// TIA Portal project "StepTimeAnalysis" (V16) (continued)
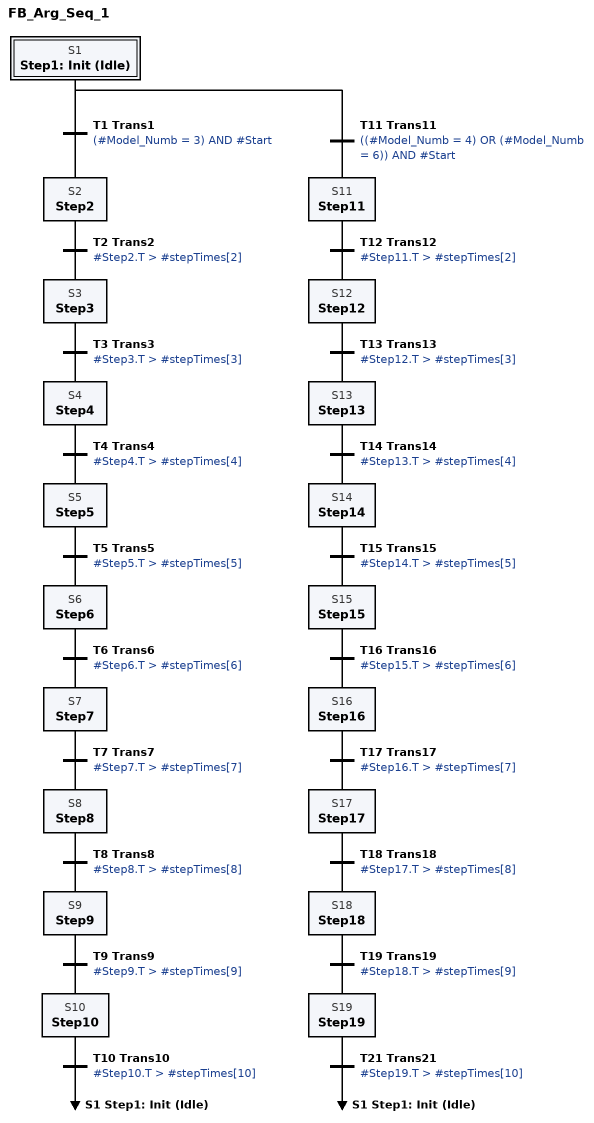
   // sequencer 1
   INITIAL_STEP "Step1: Init (Idle)":   // S1, max time T#10S, warning time T#7S
   END_STEP
   TRANSITION Trans1 FROM "Step1: Init (Idle)" TO Step2   // T1
      := (#Model_Numb = 3) AND #Start;
   END_TRANSITION
   TRANSITION Trans11 FROM "Step1: Init (Idle)" TO Step11   // T11
      := ((#Model_Numb = 4) OR (#Model_Numb = 6)) AND #Start;
   END_TRANSITION
   STEP Step2:   // S2, max time T#10S, warning time T#7S
   END_STEP
   TRANSITION Trans2 FROM Step2 TO Step3   // T2
      := #Step2.T > #stepTimes[2];
   END_TRANSITION
   STEP Step3:   // S3, max time T#10S, warning time T#7S
   END_STEP
   TRANSITION Trans3 FROM Step3 TO Step4   // T3
      := #Step3.T > #stepTimes[3];
   END_TRANSITION
   STEP Step4:   // S4, max time T#10S, warning time T#7S
   END_STEP
   TRANSITION Trans4 FROM Step4 TO Step5   // T4
      := #Step4.T > #stepTimes[4];
   END_TRANSITION
   STEP Step5:   // S5, max time T#10S, warning time T#7S
   END_STEP
   TRANSITION Trans5 FROM Step5 TO Step6   // T5
      := #Step5.T > #stepTimes[5];
   END_TRANSITION
   STEP Step6:   // S6, max time T#10S, warning time T#7S
   END_STEP
   TRANSITION Trans6 FROM Step6 TO Step7   // T6
      := #Step6.T > #stepTimes[6];
   END_TRANSITION
   STEP Step7:   // S7, max time T#10S, warning time T#7S
   END_STEP
   TRANSITION Trans7 FROM Step7 TO Step8   // T7
      := #Step7.T > #stepTimes[7];
   END_TRANSITION
   STEP Step8:   // S8, max time T#10S, warning time T#7S
   END_STEP
   TRANSITION Trans8 FROM Step8 TO Step9   // T8
      := #Step8.T > #stepTimes[8];
   END_TRANSITION
   STEP Step9:   // S9, max time T#10S, warning time T#7S
   END_STEP
   TRANSITION Trans9 FROM Step9 TO Step10   // T9
      := #Step9.T > #stepTimes[9];
   END_TRANSITION
   STEP Step10:   // S10, max time T#10S, warning time T#7S
   END_STEP
   TRANSITION Trans10 FROM Step10 TO "Step1: Init (Idle)"   // T10, jump
      := #Step10.T > #stepTimes[10];
   END_TRANSITION
   STEP Step11:   // S11, max time T#10S, warning time T#7S
   END_STEP
   TRANSITION Trans12 FROM Step11 TO Step12   // T12
      := #Step11.T > #stepTimes[2];
   END_TRANSITION
   STEP Step12:   // S12, max time T#10S, warning time T#7S
   END_STEP
   TRANSITION Trans13 FROM Step12 TO Step13   // T13
      := #Step12.T > #stepTimes[3];
   END_TRANSITION
   STEP Step13:   // S13, max time T#10S, warning time T#7S
   END_STEP
   TRANSITION Trans14 FROM Step13 TO Step14   // T14
      := #Step13.T > #stepTimes[4];
   END_TRANSITION
   STEP Step14:   // S14, max time T#10S, warning time T#7S
   END_STEP
   TRANSITION Trans15 FROM Step14 TO Step15   // T15
      := #Step14.T > #stepTimes[5];
   END_TRANSITION
   STEP Step15:   // S15, max time T#10S, warning time T#7S
   END_STEP
   TRANSITION Trans16 FROM Step15 TO Step16   // T16
      := #Step15.T > #stepTimes[6];
   END_TRANSITION
   STEP Step16:   // S16, max time T#10S, warning time T#7S
   END_STEP
   TRANSITION Trans17 FROM Step16 TO Step17   // T17
      := #Step16.T > #stepTimes[7];
   END_TRANSITION
   STEP Step17:   // S17, max time T#10S, warning time T#7S
   END_STEP
   TRANSITION Trans18 FROM Step17 TO Step18   // T18
      := #Step17.T > #stepTimes[8];
   END_TRANSITION
   STEP Step18:   // S18, max time T#10S, warning time T#7S
   END_STEP
   TRANSITION Trans19 FROM Step18 TO Step19   // T19
      := #Step18.T > #stepTimes[9];
   END_TRANSITION
   STEP Step19:   // S19, max time T#10S, warning time T#7S
   END_STEP
   TRANSITION Trans21 FROM Step19 TO "Step1: Init (Idle)"   // T21, jump
      := #Step19.T > #stepTimes[10];
   END_TRANSITION
END_FUNCTION_BLOCK

FUNCTION "FC_ARG_1" : Void   // FC1, FBD
{ S7_Optimized_Access := 'TRUE' }
VERSION : 0.1
   VAR_OUTPUT
      Ready_new_car : Bool;
   END_VAR
   VAR_TEMP
      stepTimes : Array[2..10] of Time;
      i : Int;
      Random_Time : Time;   // Random Time between 0sec to 10sec
      Start : Bool;
      Stop : Bool;
      status1_RandFunc : Word;
      status2_RandFunc : Word;
      temp : Byte;
      error_RandFunc : Bool;
   END_VAR
   VAR CONSTANT
      sequenceNO : Int := 9;
   END_VAR
BEGIN

REGION Network 1 (SCL): Man Mode Data Handling
   IF "DB_Process_Var".Man_Mode = TRUE THEN
       "DB_Process_Var".Car_Type_Selected := "DB_HMI".dropdown_selection;
   END_IF;
END_REGION

REGION Network 2 (SCL): Auto Mode Data Handling
   IF "DB_Process_Var".Auto_Mode = TRUE THEN
       "DB_HMI".dropdown_selection := 0;
       "DB_Process_Var".Car_Type_Selected := "DB_PLC2_Receiving".ReceivingBoxForward.Type;
   END_IF;
   IF "DB_HMI".ARG1_Seq1_Cmd_Auto OR "DB_HMI".Global_Cmd_Auto THEN
       "DB_HMI".dropdown_selection := 0;
       "DB_Process_Var".Car_Type_Selected := 0;
   END_IF;
END_REGION

REGION Network 3 (SCL): Load Time Date based on Car Type
       CASE "DB_Process_Var".Car_Type_Selected OF
           3:
               "DB_Profile"."time" := "DB_Profile".time_Red;
           4:
               "DB_Profile"."time" := "DB_Profile".time_Green;
           6:
               "DB_Profile"."time" := "DB_Profile".time_Blue;
       END_CASE;
END_REGION

REGION Network 4 (SCL): Switch from selected to inProduction
   IF "IDB_Arg_Seq_1_DB".Trans1.TS = TRUE OR "IDB_Arg_Seq_1_DB".Trans11.TS = TRUE THEN
       IF "DB_Process_Var".Car_Type_Selected = 3 THEN
           "DB_Process_Var".Car_Type_inProduction := 3;
           "DB_Process_Var".Car_Type_inProduction_Text := 'Red';
           "DB_HMI".ARG1_Seq1_inProduction := 3;
       ELSIF "DB_Process_Var".Car_Type_Selected = 4 THEN
           "DB_Process_Var".Car_Type_inProduction := 4;
           "DB_Process_Var".Car_Type_inProduction_Text := 'Green';
           "DB_HMI".ARG1_Seq1_inProduction := 4;
       ELSIF "DB_Process_Var".Car_Type_Selected = 6 THEN
           "DB_Process_Var".Car_Type_inProduction := 6;
           "DB_Process_Var".Car_Type_inProduction_Text := 'Blue';
           "DB_HMI".ARG1_Seq1_inProduction := 6;
       END_IF;
   END_IF;
END_REGION

REGION Network 5 (SCL): Create Random Time Values for the selected Steps
   IF "IDB_Arg_Seq_1_DB".Trans1.TS = TRUE OR "IDB_Arg_Seq_1_DB".Trans11.TS = TRUE THEN
       FOR #i := 2 TO 10 DO
           //Red
           IF "DB_HMI".ARG1_Seq1_DelaySelect_Red[#i] = TRUE THEN;
               "DB_Sim".Delta_T_Red[#i] := "LGF_RandomRange_Dint"(minValue := 0, maxValue := 10000, error => #error_RandFunc, status => #status1_RandFunc, subfunctionStatus => #status2_RandFunc);
           ELSE
               "DB_Sim".Delta_T_Red[#i] := T#0s;
           END_IF;
           //Green
           IF "DB_HMI".ARG1_Seq1_DelaySelect_Green[#i] = TRUE THEN
               "DB_Sim".Delta_T_Green[#i] := "LGF_RandomRange_Dint"(minValue := 0, maxValue := 10000, error => #error_RandFunc, status => #status1_RandFunc, subfunctionStatus => #status2_RandFunc);
           ELSE
               "DB_Sim".Delta_T_Green[#i] := T#0s;
           END_IF;
           //Blue
           IF "DB_HMI".ARG1_Seq1_DelaySelect_Blue[#i] = TRUE THEN
               "DB_Sim".Delta_T_Blue[#i] := "LGF_RandomRange_Dint"(minValue := 0, maxValue := 10000, error => #error_RandFunc, status => #status1_RandFunc, subfunctionStatus => #status2_RandFunc);
           ELSE
               "DB_Sim".Delta_T_Blue[#i] := T#0s;
           END_IF;
       END_FOR;
   END_IF;

   IF "DB_HMI".ARG1_Seq1_Cmd_DelayReset = TRUE THEN
       FOR #i := 2 TO 10 DO
           "DB_HMI".ARG1_Seq1_DelaySelect_Red[#i] := false;
           "DB_HMI".ARG1_Seq1_DelaySelect_Green[#i] := false;
           "DB_HMI".ARG1_Seq1_DelaySelect_Blue[#i] := false;
       END_FOR;
   END_IF;
END_REGION

REGION Network 6 (SCL): Add Delay Time to Step Time
   FOR #i := 2 TO 10 DO
       IF "DB_HMI".dropdown_selection = 3 OR "DB_PLC2_Receiving".ReceivingBoxForward.Type = 3 THEN
           "DB_Process_Var".Step_Times[#i] := T_ADD(IN1 := "DB_Profile"."time"[#i], IN2 := "DB_Sim".Delta_T_Red[#i]);
       ELSIF "DB_HMI".dropdown_selection = 4 OR "DB_PLC2_Receiving".ReceivingBoxForward.Type = 4 THEN
           "DB_Process_Var".Step_Times[#i] := T_ADD(IN1 := "DB_Profile"."time"[#i], IN2 := "DB_Sim".Delta_T_Green[#i]);
       ELSIF "DB_HMI".dropdown_selection = 6 OR "DB_PLC2_Receiving".ReceivingBoxForward.Type = 6 THEN
           "DB_Process_Var".Step_Times[#i] := T_ADD(IN1 := "DB_Profile"."time"[#i], IN2 := "DB_Sim".Delta_T_Blue[#i]);
       END_IF;
   END_FOR;
END_REGION

REGION Network 7: Auto Mode select
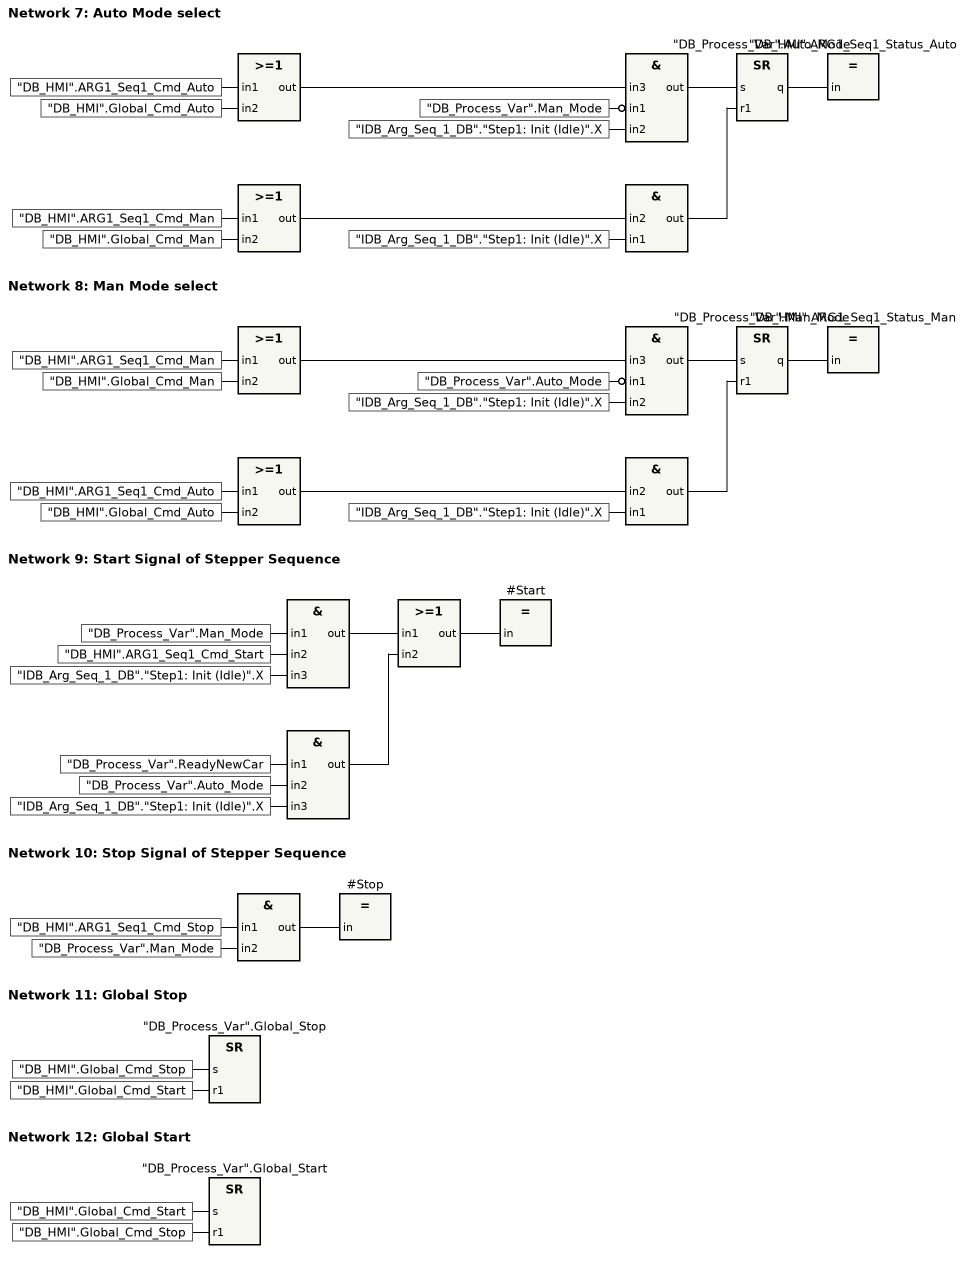
   IF ("DB_HMI".ARG1_Seq1_Cmd_Auto OR "DB_HMI".Global_Cmd_Auto) AND NOT "DB_Process_Var".Man_Mode AND "IDB_Arg_Seq_1_DB"."Step1: Init (Idle)".X THEN
       "DB_Process_Var".Auto_Mode := TRUE;   // SR flip-flop
   END_IF;
   IF ("DB_HMI".ARG1_Seq1_Cmd_Man OR "DB_HMI".Global_Cmd_Man) AND "IDB_Arg_Seq_1_DB"."Step1: Init (Idle)".X THEN
       "DB_Process_Var".Auto_Mode := FALSE;
   END_IF;
   "DB_HMI".ARG1_Seq1_Status_Auto := "DB_Process_Var".Auto_Mode;
END_REGION

REGION Network 8: Man Mode select
   IF ("DB_HMI".ARG1_Seq1_Cmd_Man OR "DB_HMI".Global_Cmd_Man) AND NOT "DB_Process_Var".Auto_Mode AND "IDB_Arg_Seq_1_DB"."Step1: Init (Idle)".X THEN
       "DB_Process_Var".Man_Mode := TRUE;   // SR flip-flop
   END_IF;
   IF ("DB_HMI".ARG1_Seq1_Cmd_Auto OR "DB_HMI".Global_Cmd_Auto) AND "IDB_Arg_Seq_1_DB"."Step1: Init (Idle)".X THEN
       "DB_Process_Var".Man_Mode := FALSE;
   END_IF;
   "DB_HMI".ARG1_Seq1_Status_Man := "DB_Process_Var".Man_Mode;
END_REGION

REGION Network 9: Start Signal of Stepper Sequence
   #Start := ("DB_Process_Var".Man_Mode AND "DB_HMI".ARG1_Seq1_Cmd_Start AND "IDB_Arg_Seq_1_DB"."Step1: Init (Idle)".X) OR ("DB_Process_Var".ReadyNewCar AND "DB_Process_Var".Auto_Mode AND "IDB_Arg_Seq_1_DB"."Step1: Init (Idle)".X);
END_REGION

REGION Network 10: Stop Signal of Stepper Sequence
   #Stop := "DB_HMI".ARG1_Seq1_Cmd_Stop AND "DB_Process_Var".Man_Mode;
END_REGION

REGION Network 11: Global Stop
   IF "DB_HMI".Global_Cmd_Stop THEN
       "DB_Process_Var".Global_Stop := TRUE;   // SR flip-flop
   END_IF;
   IF "DB_HMI".Global_Cmd_Start THEN "DB_Process_Var".Global_Stop := FALSE; END_IF;
END_REGION

REGION Network 12: Global Start
   IF "DB_HMI".Global_Cmd_Start THEN
       "DB_Process_Var".Global_Start := TRUE;   // SR flip-flop
   END_IF;
   IF "DB_HMI".Global_Cmd_Stop THEN "DB_Process_Var".Global_Start := FALSE; END_IF;
END_REGION

REGION Network 13 (SCL): Reset Type Selection
   IF "DB_HMI".ARG1_Seq1_Cmd_Stop = TRUE THEN
       "DB_PLC2_Receiving".ReceivingBoxForward.Type := 0;
       "DB_HMI".ARG1_Seq1_inProduction := 0;
       "DB_Process_Var".ReadyNewCar := TRUE;
   END_IF;
END_REGION

REGION Network 14: Call FB with Stepper Sequence
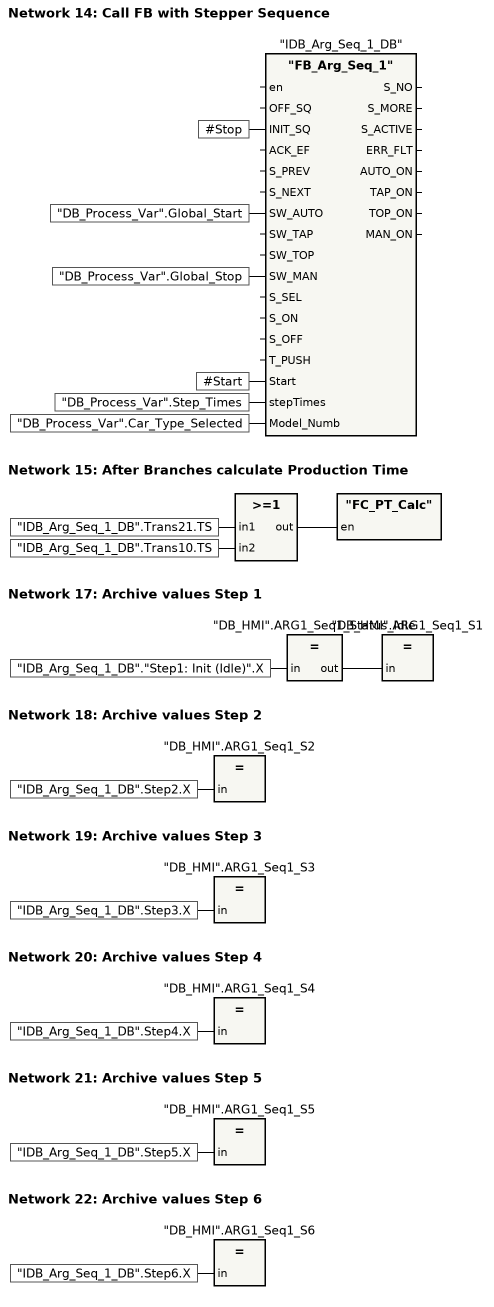
   "IDB_Arg_Seq_1_DB"(INIT_SQ := #Stop,   // "FB_Arg_Seq_1"
                      SW_AUTO := "DB_Process_Var".Global_Start,
                      SW_MAN := "DB_Process_Var".Global_Stop,
                      Start := #Start,
                      stepTimes := "DB_Process_Var".Step_Times,
                      Model_Numb := "DB_Process_Var".Car_Type_Selected);
END_REGION

REGION Network 15: After Branches calculate Production Time
   IF "IDB_Arg_Seq_1_DB".Trans21.TS OR "IDB_Arg_Seq_1_DB".Trans10.TS THEN "FC_PT_Calc"(); END_IF;
END_REGION

REGION Network 16 (SCL): Send Idle to previous Station
   IF "IDB_Arg_Seq_1_DB"."Step1: Init (Idle)".X = TRUE THEN
       "DB_PLC2_Sending".SendBox.Station_Idle := TRUE;
   ELSE
       "DB_PLC2_Sending".SendBox.Station_Idle := FALSE;
   END_IF;
END_REGION

REGION Network 17: Archive values Step 1
   "DB_HMI".ARG1_Seq1_Status_Idle := "IDB_Arg_Seq_1_DB"."Step1: Init (Idle)".X;
   "DB_HMI".ARG1_Seq1_S1 := "IDB_Arg_Seq_1_DB"."Step1: Init (Idle)".X;
END_REGION

REGION Network 18: Archive values Step 2
   "DB_HMI".ARG1_Seq1_S2 := "IDB_Arg_Seq_1_DB".Step2.X;
END_REGION

REGION Network 19: Archive values Step 3
   "DB_HMI".ARG1_Seq1_S3 := "IDB_Arg_Seq_1_DB".Step3.X;
END_REGION

REGION Network 20: Archive values Step 4
   "DB_HMI".ARG1_Seq1_S4 := "IDB_Arg_Seq_1_DB".Step4.X;
END_REGION

REGION Network 21: Archive values Step 5
   "DB_HMI".ARG1_Seq1_S5 := "IDB_Arg_Seq_1_DB".Step5.X;
END_REGION

REGION Network 22: Archive values Step 6
   "DB_HMI".ARG1_Seq1_S6 := "IDB_Arg_Seq_1_DB".Step6.X;
END_REGION

REGION Network 23: Archive values Step 7
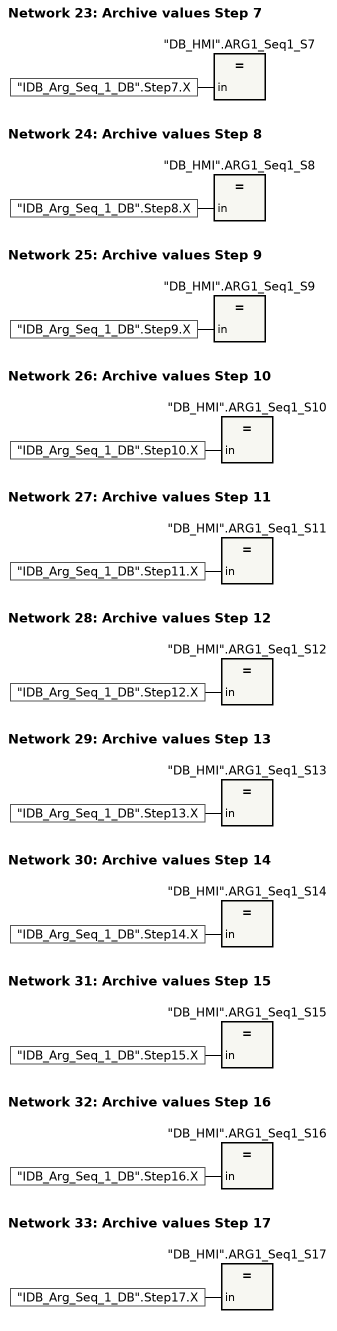
   "DB_HMI".ARG1_Seq1_S7 := "IDB_Arg_Seq_1_DB".Step7.X;
END_REGION

REGION Network 24: Archive values Step 8
   "DB_HMI".ARG1_Seq1_S8 := "IDB_Arg_Seq_1_DB".Step8.X;
END_REGION

REGION Network 25: Archive values Step 9
   "DB_HMI".ARG1_Seq1_S9 := "IDB_Arg_Seq_1_DB".Step9.X;
END_REGION

REGION Network 26: Archive values Step 10
   "DB_HMI".ARG1_Seq1_S10 := "IDB_Arg_Seq_1_DB".Step10.X;
END_REGION

REGION Network 27: Archive values Step 11
   "DB_HMI".ARG1_Seq1_S11 := "IDB_Arg_Seq_1_DB".Step11.X;
END_REGION

REGION Network 28: Archive values Step 12
   "DB_HMI".ARG1_Seq1_S12 := "IDB_Arg_Seq_1_DB".Step12.X;
END_REGION

REGION Network 29: Archive values Step 13
   "DB_HMI".ARG1_Seq1_S13 := "IDB_Arg_Seq_1_DB".Step13.X;
END_REGION

REGION Network 30: Archive values Step 14
   "DB_HMI".ARG1_Seq1_S14 := "IDB_Arg_Seq_1_DB".Step14.X;
END_REGION

REGION Network 31: Archive values Step 15
   "DB_HMI".ARG1_Seq1_S15 := "IDB_Arg_Seq_1_DB".Step15.X;
END_REGION

REGION Network 32: Archive values Step 16
   "DB_HMI".ARG1_Seq1_S16 := "IDB_Arg_Seq_1_DB".Step16.X;
END_REGION

REGION Network 33: Archive values Step 17
   "DB_HMI".ARG1_Seq1_S17 := "IDB_Arg_Seq_1_DB".Step17.X;
END_REGION

REGION Network 34: Archive values Step 18
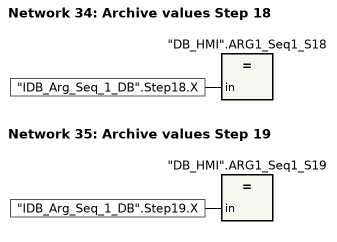
   "DB_HMI".ARG1_Seq1_S18 := "IDB_Arg_Seq_1_DB".Step18.X;
END_REGION

REGION Network 35: Archive values Step 19
   "DB_HMI".ARG1_Seq1_S19 := "IDB_Arg_Seq_1_DB".Step19.X;
END_REGION

REGION Network 36 (SCL): Set Busy
   IF
       "IDB_Arg_Seq_1_DB".Step2.X OR
       "IDB_Arg_Seq_1_DB".Step3.X OR
       "IDB_Arg_Seq_1_DB".Step4.X OR
       "IDB_Arg_Seq_1_DB".Step5.X OR
       "IDB_Arg_Seq_1_DB".Step6.X OR
       "IDB_Arg_Seq_1_DB".Step7.X OR
       "IDB_Arg_Seq_1_DB".Step8.X OR
       "IDB_Arg_Seq_1_DB".Step9.X OR
       "IDB_Arg_Seq_1_DB".Step10.X OR
       "IDB_Arg_Seq_1_DB".Step11.X OR
       "IDB_Arg_Seq_1_DB".Step12.X OR
       "IDB_Arg_Seq_1_DB".Step13.X OR
       "IDB_Arg_Seq_1_DB".Step14.X OR
       "IDB_Arg_Seq_1_DB".Step15.X OR
       "IDB_Arg_Seq_1_DB".Step16.X OR
       "IDB_Arg_Seq_1_DB".Step17.X OR
       "IDB_Arg_Seq_1_DB".Step18.X OR
       "IDB_Arg_Seq_1_DB".Step19.X THEN
       "DB_HMI".ARG1_Seq1_Status_Busy := TRUE;
   ELSIF "IDB_Arg_Seq_1_DB"."Step1: Init (Idle)".X THEN
       "DB_HMI".ARG1_Seq1_Status_Busy := FALSE;
   END_IF;
END_REGION

REGION Network 37 (SCL): When Stepper Sequence runs completely
   IF "IDB_Arg_Seq_1_DB".Trans10.TS = TRUE OR "IDB_Arg_Seq_1_DB".Trans21.TS = TRUE THEN
       "DB_Process_Var".Branch_Complete := TRUE;
       "DB_Process_Var".Car_Type_Ready := "DB_Process_Var".Car_Type_inProduction;
       "DB_Process_Var".Car_Type_inProduction := 0;
       "DB_Process_Var".Car_Type_inProduction_Text := '';
       "DB_Process_Var".Car_ReadyToShift := TRUE;
       "DB_HMI".ARG1_Seq1_inProduction := 0;
   END_IF;
   IF "IDB_Arg_Seq_1_DB".Trans1.TS = TRUE OR "IDB_Arg_Seq_1_DB".Trans11.TS = TRUE THEN
       "DB_Process_Var".Branch_Complete := FALSE;
       "DB_Process_Var".ReadyNewCar := 0;
   END_IF;
END_REGION

REGION Network 38 (SCL): Write Data in the Sending Box
   //IF "DB_Process_Var".Branch_Complete = TRUE AND "DB_PLC2_Receiving".ReceivingBox.Station_Idle = TRUE THEN
   IF "IDB_Arg_Seq_1_DB".Trans10.TS = TRUE OR "IDB_Arg_Seq_1_DB".Trans21.TS = TRUE THEN
       "DB_PLC2_Sending".SendBoxForward.Planned_PT_Red := "DB_HMI".ARG1_Seq1_Calculated_PT_Red;
       "DB_PLC2_Sending".SendBoxForward.Planned_PT_Green := "DB_HMI".ARG1_Seq1_Calculated_PT_Green;
       "DB_PLC2_Sending".SendBoxForward.Planned_PT_Blue := "DB_HMI".ARG1_Seq1_Calculated_PT_Blue;

       "DB_PLC2_Sending".SendBoxForward.Measuered_PT_Red := "DB_HMI".ARG1_Seq1_Messured_PT_Red;
       "DB_PLC2_Sending".SendBoxForward.Measuered_PT_Green := "DB_HMI".ARG1_Seq1_Messured_PT_Green;
       "DB_PLC2_Sending".SendBoxForward.Measuered_PT_Blue := "DB_HMI".ARG1_Seq1_Messured_PT_Blue;

       "DB_PLC2_Sending".SendBoxForward.Type := "DB_Process_Var".Car_Type_Ready;

       "DB_PLC2_Receiving".ReceivingBoxForward.Type := 0;
   END_IF;
END_REGION

REGION Network 39 (SCL): Reset Receiving Car Typ
   //IF "IDB_Arg_Seq_1_DB".Trans1.TS = TRUE OR "IDB_Arg_Seq_1_DB".Trans11.TS THEN
       //"DB_PLC2_Receiving".ReceivingBoxForward.Type := 0;
   //END_IF;
END_REGION

REGION Network 40 (SCL): When car is shifted
   IF "DB_Process_Var".Data_Put_Done = TRUE THEN
       "DB_Process_Var".Car_Type_Ready := 0;
       "DB_PLC2_Sending".SendBoxForward.Type := 0;
       "DB_Process_Var".Car_ReadyToShift := FALSE;
       "DB_HMI".ARG1_Seq1_inProduction := 0;
       "DB_Process_Var".ReadyNewCar := 1;

       //"DB_PLC2_Receiving".ReceivingBoxForward.Type := 0;
   END_IF;
END_REGION
END_FUNCTION

FUNCTION "FC_Com" : Void   // FC2, FBD
{ S7_Optimized_Access := 'TRUE' }
VERSION : 0.1
BEGIN

REGION Network 1: Communication PLC1 -> PLC2
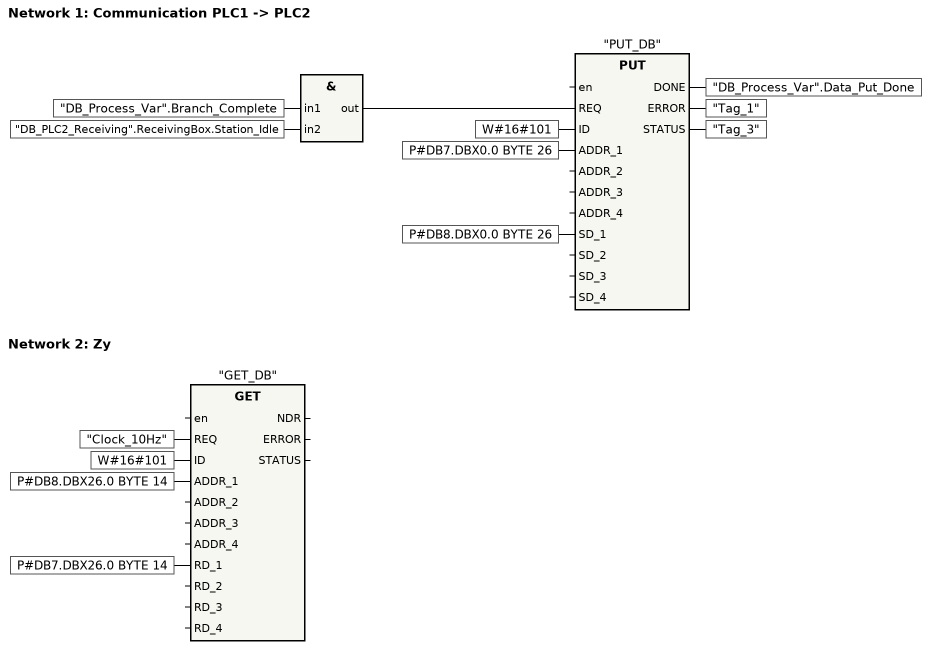
   "PUT_DB"(REQ := "DB_Process_Var".Branch_Complete AND "DB_PLC2_Receiving".ReceivingBox.Station_Idle,   // PUT
            ID := W#16#101,
            ADDR_1 := P#DB7.DBX0.0 BYTE 26,
            SD_1 := P#DB8.DBX0.0 BYTE 26,
            DONE => "DB_Process_Var".Data_Put_Done,
            ERROR => "Tag_1",
            STATUS => "Tag_3");
END_REGION

REGION Network 2: Zy
   "GET_DB"(REQ := "Clock_10Hz", ID := W#16#101, ADDR_1 := P#DB8.DBX26.0 BYTE 14, RD_1 := P#DB7.DBX26.0 BYTE 14);   // GET
END_REGION
END_FUNCTION

FUNCTION "FC_PT_Calc" : Void   // FC3, SCL
{ S7_Optimized_Access := 'TRUE' }
VERSION : 0.1
   VAR_TEMP
      i : Int;
   END_VAR
   VAR CONSTANT
      sequenceNO : Int := 9;
      Null : Time := T#0MS;
   END_VAR
BEGIN
   "DB_HMI".ARG1_Seq1_Calculated_PT_Red := #Null;
   "DB_HMI".ARG1_Seq1_Calculated_PT_Green := #Null;
   "DB_HMI".ARG1_Seq1_Calculated_PT_Blue := #Null;

   "DB_HMI".ARG1_Seq1_Messured_PT_Red := #Null;
   "DB_HMI".ARG1_Seq1_Messured_PT_Green := #Null;
   "DB_HMI".ARG1_Seq1_Messured_PT_Blue := #Null;

   FOR #i := 2 TO #sequenceNO + 1 DO
       //Calculated Production Time
       "DB_HMI".ARG1_Seq1_Calculated_PT_Red := "DB_HMI".ARG1_Seq1_Calculated_PT_Red + "DB_Profile".time_Red[#i];
       "DB_HMI".ARG1_Seq1_Calculated_PT_Green := "DB_HMI".ARG1_Seq1_Calculated_PT_Green + "DB_Profile".time_Green[#i];
       "DB_HMI".ARG1_Seq1_Calculated_PT_Blue := "DB_HMI".ARG1_Seq1_Calculated_PT_Blue + "DB_Profile".time_Blue[#i];
       //Messured Production Time
       IF "DB_Process_Var".Car_Type_inProduction = 3 THEN
           "DB_HMI".ARG1_Seq1_Messured_PT_Red := "DB_HMI".ARG1_Seq1_Messured_PT_Red + "DB_Process_Var".Step_Times[#i];
       ELSIF "DB_Process_Var".Car_Type_inProduction = 4 THEN
           "DB_HMI".ARG1_Seq1_Messured_PT_Green := "DB_HMI".ARG1_Seq1_Messured_PT_Green + "DB_Process_Var".Step_Times[#i];
       ELSIF "DB_Process_Var".Car_Type_inProduction = 6 THEN
           "DB_HMI".ARG1_Seq1_Messured_PT_Blue := "DB_HMI".ARG1_Seq1_Messured_PT_Blue + "DB_Process_Var".Step_Times[#i];
       END_IF;
   END_FOR;

   //Add Time of previous Stations
   "DB_HMI".ARG1_Seq1_Calculated_PT_Red := "DB_HMI".ARG1_Seq1_Calculated_PT_Red + "DB_PLC2_Receiving".ReceivingBoxForward.Planned_PT_Red;
   "DB_HMI".ARG1_Seq1_Calculated_PT_Green := "DB_HMI".ARG1_Seq1_Calculated_PT_Green + "DB_PLC2_Receiving".ReceivingBoxForward.Planned_PT_Green;
   "DB_HMI".ARG1_Seq1_Calculated_PT_Blue := "DB_HMI".ARG1_Seq1_Calculated_PT_Blue + "DB_PLC2_Receiving".ReceivingBoxForward.Planned_PT_Blue;

   "DB_HMI".ARG1_Seq1_Messured_PT_Red := "DB_HMI".ARG1_Seq1_Messured_PT_Red + "DB_PLC2_Receiving".ReceivingBoxForward.Measuered_PT_Red;
   "DB_HMI".ARG1_Seq1_Messured_PT_Green := "DB_HMI".ARG1_Seq1_Messured_PT_Green + "DB_PLC2_Receiving".ReceivingBoxForward.Measuered_PT_Green;
   "DB_HMI".ARG1_Seq1_Messured_PT_Blue := "DB_HMI".ARG1_Seq1_Messured_PT_Blue + "DB_PLC2_Receiving".ReceivingBoxForward.Measuered_PT_Blue;
END_FUNCTION

FUNCTION "FC_Global_Status" : Void   // FC4, SCL
{ S7_Optimized_Access := 'TRUE' }
VERSION : 0.1
   VAR_TEMP
      global_auto : Bool;
      global_man : Bool;
   END_VAR
BEGIN
   IF "DB_Process_Var".Auto_Mode = TRUE THEN
       "DB_PLC2_Sending".SendBox.Mode_PLC2 := 1;
   ELSIF "DB_Process_Var".Man_Mode = TRUE THEN
       "DB_PLC2_Sending".SendBox.Mode_PLC2 := 2;
   ELSE
       "DB_PLC2_Sending".SendBox.Mode_PLC2 := 0;
   END_IF;

   "DB_PLC2_Sending".SendBox.Mode_PLC5 := "DB_PLC2_Receiving".ReceivingBox.Mode_PLC5;
   "DB_PLC2_Sending".SendBox.Mode_PLC4 := "DB_PLC2_Receiving".ReceivingBox.Mode_PLC4;
   "DB_PLC2_Sending".SendBox.Mode_PLC3 := "DB_PLC2_Receiving".ReceivingBox.Mode_PLC3;

   IF "DB_Process_Var".Station_Nr = 1 THEN
       IF "DB_PLC2_Sending".SendBox.Mode_PLC2 = 1 AND "DB_PLC2_Receiving".ReceivingBox.Mode_PLC2 = 1 AND "DB_PLC2_Receiving".ReceivingBox.Mode_PLC3 = 1 AND "DB_PLC2_Receiving".ReceivingBox.Mode_PLC4 = 1 AND "DB_PLC2_Receiving".ReceivingBox.Mode_PLC5 = 1 THEN
           "DB_HMI".Global_Status_Auto := TRUE;
       ELSIF "DB_PLC2_Sending".SendBox.Mode_PLC2 = 0 AND "DB_PLC2_Receiving".ReceivingBox.Mode_PLC2 = 0 AND "DB_PLC2_Receiving".ReceivingBox.Mode_PLC3 = 0 AND "DB_PLC2_Receiving".ReceivingBox.Mode_PLC4 = 0 AND "DB_PLC2_Receiving".ReceivingBox.Mode_PLC5 = 0 THEN
           "DB_HMI".Global_Status_Auto := FALSE;
           "DB_HMI".Global_Status_Man := FALSE;
       ELSE
           "DB_HMI".Global_Status_Man := TRUE;
       END_IF;
   END_IF;
END_FUNCTION

ORGANIZATION_BLOCK "Main"   // OB1, LAD, ProgramCycle
TITLE = "Main Program Sweep (Cycle)"
{ S7_Optimized_Access := 'TRUE' }
VERSION : 0.1
   VAR_INPUT
      Initial_Call : Bool;   // Initial call of this OB
      Remanence : Bool;   // =True, if remanent data are available
   END_VAR
   VAR_TEMP
      test : Bool;
   END_VAR
BEGIN

REGION Network 1: Call ARG_1
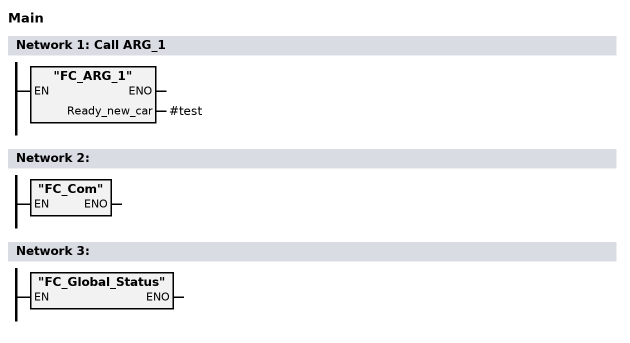
   RUNG wire#powerrail
      "FC_ARG_1"(Ready_new_car => #test)
   END_RUNG
   // the same network as SCL:
   "FC_ARG_1"(Ready_new_car => #test);
END_REGION

REGION Network 2
   RUNG wire#powerrail
      "FC_Com"()
   END_RUNG
   // the same network as SCL:
   "FC_Com"();
END_REGION

REGION Network 3
   RUNG wire#powerrail
      "FC_Global_Status"()
   END_RUNG
   // the same network as SCL:
   "FC_Global_Status"();
END_REGION
END_ORGANIZATION_BLOCK

// folder: LGF/4 Math operations

FUNCTION "LGF_RandomRange_Dint" : DInt   // FC10013, SCL
TITLE = LGF_RandomRange_DInt
{ S7_Optimized_Access := 'TRUE' }
AUTHOR : Siemens_Digital_Industries
FAMILY : LGF
NAME : LGF_RandomRange_DInt
// This function generates random numbers in defined limits (Datatype DInt)
   VAR_INPUT
      minValue : DInt;   // minimal Value random can reach / Minimum value of the range of the random number
      maxValue : DInt;   // maximal Value random can reach / Maximum value of the range of the random number
   END_VAR
   VAR_OUTPUT
      error : Bool;   // Error if true
      status : Word;   // Status of the function
      subfunctionStatus : Word;   // Status or return value of called FB's, FCs and system blocks
   END_VAR
   VAR_TEMP
      tempTime : DTL;   // System time
      tempNanoSecondInDWord : DWord;   // UDINT converted to DWORD for access to individual bytes
      tempTimeStatus : Word;   // Status of the instruction RD_SYS_T
      tempRandomValue : DWord;   // Random-start-value
      tempNormReal : Real;   // Normalized value
   END_VAR
   // Ret_Val : Returns random DInt number in a predefined range
   VAR CONSTANT
      ZERO : DInt := 0;   // Zero value in case of error
      MAX_UDINT : UDInt := 4294967295 ;   // Maximum UDINT value
      SUB_STATUS_NO_ERROR : Word := 16#0000;   // Status: sub function call ends without error
      STATUS_FINISHED_NO_ERROR : Word := 16#0000;   // Status: Execution finished without errors
      ERR_MAX_LESS_MIN : Word := 16#8200;   // Error: The maximum limit number is smaller than the minimum limit number
      ERR_RD_SYS_T : Word := 16#8600;   // Error: System function Read system time returned an error
   END_VAR
BEGIN
   REGION Block info header
     //=============================================================================
     // SIEMENS AG / (c)Copyright 2017
     //-----------------------------------------------------------------------------
     // Title:            LGF_RandomRange_DInt
     // Comment/Function: This function generates random numbers in defined limits (Datatype DInt)
     // Library/Family:   LGF(Library General Functions)
     // Author:           Siemens Digital Industry Support
     // Tested with:      S7-PLCSIM Advanced V2.0 SP1
     // Engineering:      TIA Portal V15 Update 2
     // Restrictions:     ENO disabled - error handling done by error and status
     // Requirements:     PLC (S7-1200 / S7-1500)
     //-------------------------------------------------------------------------------
     // Change log table:
     // Version  | Date       | Expert in charge       | Changes applied
     //----------|------------|------------------------|------------------------------
     // 01.00.00 19.08.2015  Siemens Industry Online Support
     //                      First released version
     // 01.00.01 02.01.2017  Siemens Industry Online Support
     //                      Upgrade: TIA Portal V14 Update 1
     // 01.00.02 17.08.2018  Siemens Industry Online Support
     //                      Upgrade: TIA V15 Update 2
     // 01.00.03 23.11.2018  Siemens Industry Online Support
     //                      Upgrade: TIA V15.1
     // 01.01.00 09.10.2019  Siemens Industry Presales Support
     //                      Renamed from "LGF_RandomInt" to "LGF_RandomRange_DInt"
     //                      change random datatype from int to dint
     //                      Regions, commens and costants are added
     // 03.00.00 23.04.2020  Siemens Industry Support
     //                      Set version to V3.0.0, harmonize the version of the whole library
     //=============================================================================
   END_REGION

   REGION Validation
     // Check if the maximal Value is less than the minimal value
     IF (#minValue > #maxValue) THEN
       #error := true;
       #status := #ERR_MAX_LESS_MIN;
       #subfunctionStatus := #SUB_STATUS_NO_ERROR;
       #LGF_RandomRange_Dint := #ZERO;
       RETURN;
     END_IF;

     // Read system time
     #tempTimeStatus := INT_TO_WORD(RD_SYS_T(#tempTime));

     // Check return variable for error
     IF (#tempTimeStatus <> #SUB_STATUS_NO_ERROR) THEN
       #error := true;
       #status := #ERR_RD_SYS_T;
       #subfunctionStatus := #tempTimeStatus;
       #LGF_RandomRange_Dint := #ZERO;
       RETURN;
     END_IF;
   END_REGION

   REGION Calculating random number
     // Converting to double word so individual bytes can be addressed
     #tempNanoSecondInDWord := UDINT_TO_DWORD(#tempTime.NANOSECOND);

     // Callculate a random-start-value depending on the time
     #tempRandomValue.%B3 := #tempNanoSecondInDWord.%B0;
     #tempRandomValue.%B2 := #tempNanoSecondInDWord.%B1;
     #tempRandomValue.%B1 := #tempNanoSecondInDWord.%B2;
     #tempRandomValue.%B0 := #tempNanoSecondInDWord.%B3;

     // Norm the calculated random number: 0.0 <= #tempNormReal <= 1.0
     #tempNormReal := UDINT_TO_REAL(DWORD_TO_UDINT(#tempRandomValue)) / UDINT_TO_REAL(#MAX_UDINT);

     // Scale the tempNormReal to be in the range of maxValue and minValue
     #LGF_RandomRange_Dint := REAL_TO_DINT((#tempNormReal * DINT_TO_REAL(#maxValue - #minValue) + DINT_TO_REAL(#minValue)));

     #error := false;
     #status := #STATUS_FINISHED_NO_ERROR;
     #subfunctionStatus := #SUB_STATUS_NO_ERROR;
     // ENO mechanism is not used
     ENO := TRUE;
   END_REGION
END_FUNCTION

FUNCTION "LGF_Random_DInt" : DInt   // FC10084, SCL
TITLE = LGF_Random_DInt
{ S7_Optimized_Access := 'TRUE' }
AUTHOR : Siemens_Digital_Industries
FAMILY : LGF
NAME : LGF_Random_DInt
// Generates a random number in the DInt Range
   VAR_OUTPUT
      error : Bool;   // Error if true
      status : Word;   // Status of the function
      subfunctionStatus : Word;   // Status or return value of called FB's, FCs and system blocks
   END_VAR
   VAR_TEMP
      tempTime : DTL;   // System time
      tempNanoSecondInDWord : DWord;   // UDINT converted to DWORD for access to individual bytes
      tempTimeStatus : Word;   // Status of the instruction RD_SYS_T
      tempRandomValue : DWord;   // Random-start-value
   END_VAR
   // Ret_Val : Random number in the Dint range
   VAR CONSTANT
      ZERO : DInt;   // Zero value in case of error
      SUB_STATUS_NO_ERROR : Word := 16#0000;   // Status: sub function call ends without error
      STATUS_FINISHED_NO_ERROR : Word := 16#0000;   // Status: Execution finished without errors
      ERR_RD_SYS_T : Word := 16#8600;   // Error: System function Read system time returned an error
   END_VAR
BEGIN
   REGION Block info header
     //=============================================================================
     // SIEMENS AG / (c)Copyright 2017
     //-----------------------------------------------------------------------------
     // Title:            LGF_Random_DInt
     // Comment/Function: Generates a random number in the DInt Range
     // Library/Family:   LGF(Library General Functions)
     // Author:           Siemens Digital Industry Support
     // Tested with:      S7-PLCSIM Advanced V2.0 SP1
     // Engineering:      TIA Portal V15 Update 2
     // Restrictions:     ENO disabled - error handling done by error and status
     // Requirements:     PLC (S7-1200 / S7-1500)
     //-------------------------------------------------------------------------------
     // Change log table:
     // Version  | Date       | Expert in charge       | Changes applied
     //----------|------------|------------------------|------------------------------
     // 01.00.00 13.11.2019  Siemens Industry Presales Support
     //                      First release
     //                      copied from "LGF_Random_Real"
     // 03.00.00 23.04.2020  Siemens Industry Support
     //                      Set version to V3.0.0, harmonize the version of the whole library
     //=============================================================================
   END_REGION

   REGION Validation
     // Read system time
     #tempTimeStatus := INT_TO_WORD(RD_SYS_T(#tempTime));

     // Check return variable for error
     IF (#tempTimeStatus <> #SUB_STATUS_NO_ERROR) THEN
       #error := true;
       #status := #ERR_RD_SYS_T;
       #subfunctionStatus := #tempTimeStatus;
       #LGF_Random_DInt := #ZERO;
       RETURN;
     END_IF;
   END_REGION

   REGION Calculating random number
     // Converting to double word so individual bytes can be addressed
     #tempNanoSecondInDWord := UDINT_TO_DWORD(#tempTime.NANOSECOND);

     // Calculate a random-start-value depending on the time
     #tempRandomValue.%B3 := #tempNanoSecondInDWord.%B0;
     #tempRandomValue.%B2 := #tempNanoSecondInDWord.%B1;
     #tempRandomValue.%B1 := #tempNanoSecondInDWord.%B2;
     #tempRandomValue.%B0 := #tempNanoSecondInDWord.%B3;

     #LGF_Random_DInt := DWORD_TO_DINT(#tempRandomValue);

     #error := false;
     #status := #STATUS_FINISHED_NO_ERROR;
     #subfunctionStatus := #SUB_STATUS_NO_ERROR;
     // ENO mechanism is not used
     ENO := TRUE;
   END_REGION
END_FUNCTION

// ===== PLC "PLC_3"  CPU 1517TF-3 PN/DP =====

VAR_GLOBAL   // PLC tag table "Standard-Variablentabelle"
   "Clock_Byte" AT %MB0 : Byte;
   "Clock_10Hz" AT %M0.0 : Bool;
   "Clock_5Hz" AT %M0.1 : Bool;
   "Clock_2.5Hz" AT %M0.2 : Bool;
   "Clock_2Hz" AT %M0.3 : Bool;
   "Clock_1.25Hz" AT %M0.4 : Bool;
   "Clock_1Hz" AT %M0.5 : Bool;
   "Clock_0.625Hz" AT %M0.6 : Bool;
   "Clock_0.5Hz" AT %M0.7 : Bool;
   "Tag_1" AT %M10.1 : Bool;
   "Tag_2" AT %M10.2 : Bool;
   "Tag_3" AT %MW14 : Word;
END_VAR

TYPE "PLC_SF"
   STRUCT
      "Type" : Int;
      Planned_PT_Red : Time;
      Planned_PT_Green : Time;
      Planned_PT_Blue : Time;
      Measuered_PT_Red : Time;
      Measuered_PT_Green : Time;
      Measuered_PT_Blue : Time;
   END_STRUCT;
END_TYPE

TYPE "PLC_SR"
   STRUCT
      "Type" : Int;
      Station_Idle : Bool;
      Mode_PLC1 : Int;
      Mode_PLC2 : Int;
      Mode_PLC3 : Int;
      Mode_PLC4 : Int;
      Mode_PLC5 : Int;
   END_STRUCT;
END_TYPE

DATA_BLOCK "IDB_Arg_Seq_1_DB"   // DB2
{ S7_Optimized_Access := 'TRUE' }
VERSION : 0.1
// stored: InstanceOfName FB_Arg_Seq_1
"FB_Arg_Seq_1"
BEGIN
END_DATA_BLOCK

